REGION Network 15: EM - Abort Command
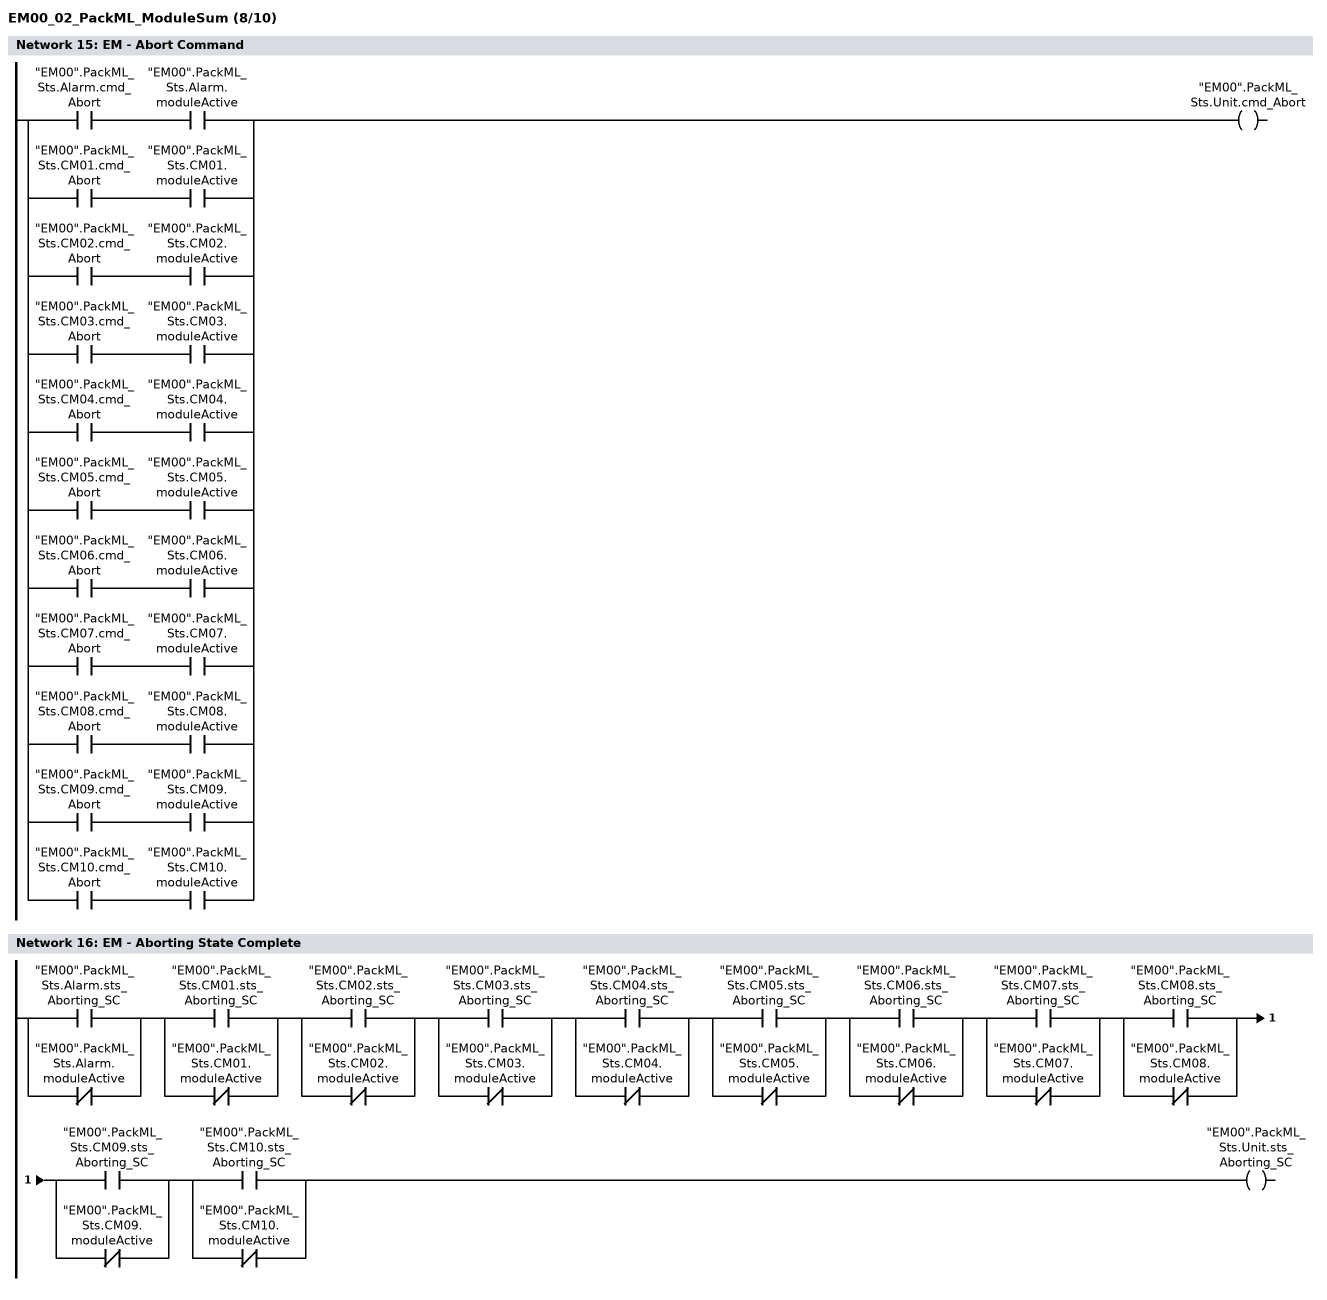
   RUNG wire#powerrail
      Contact( "EM00".PackML_Sts.Alarm.cmd_Abort )
      Contact( "EM00".PackML_Sts.Alarm.moduleActive )
      wire#w1
      Coil( "EM00".PackML_Sts.Unit.cmd_Abort )
   END_RUNG
   RUNG wire#powerrail
      Contact( "EM00".PackML_Sts.CM01.cmd_Abort )
      Contact( "EM00".PackML_Sts.CM01.moduleActive )
   END_RUNG wire#w1
   RUNG wire#powerrail
      Contact( "EM00".PackML_Sts.CM02.cmd_Abort )
      Contact( "EM00".PackML_Sts.CM02.moduleActive )
   END_RUNG wire#w1
   RUNG wire#powerrail
      Contact( "EM00".PackML_Sts.CM03.cmd_Abort )
      Contact( "EM00".PackML_Sts.CM03.moduleActive )
   END_RUNG wire#w1
   RUNG wire#powerrail
      Contact( "EM00".PackML_Sts.CM04.cmd_Abort )
      Contact( "EM00".PackML_Sts.CM04.moduleActive )
   END_RUNG wire#w1
   RUNG wire#powerrail
      Contact( "EM00".PackML_Sts.CM05.cmd_Abort )
      Contact( "EM00".PackML_Sts.CM05.moduleActive )
   END_RUNG wire#w1
   RUNG wire#powerrail
      Contact( "EM00".PackML_Sts.CM06.cmd_Abort )
      Contact( "EM00".PackML_Sts.CM06.moduleActive )
   END_RUNG wire#w1
   RUNG wire#powerrail
      Contact( "EM00".PackML_Sts.CM07.cmd_Abort )
      Contact( "EM00".PackML_Sts.CM07.moduleActive )
   END_RUNG wire#w1
   RUNG wire#powerrail
      Contact( "EM00".PackML_Sts.CM08.cmd_Abort )
      Contact( "EM00".PackML_Sts.CM08.moduleActive )
   END_RUNG wire#w1
   RUNG wire#powerrail
      Contact( "EM00".PackML_Sts.CM09.cmd_Abort )
      Contact( "EM00".PackML_Sts.CM09.moduleActive )
   END_RUNG wire#w1
   RUNG wire#powerrail
      Contact( "EM00".PackML_Sts.CM10.cmd_Abort )
      Contact( "EM00".PackML_Sts.CM10.moduleActive )
   END_RUNG wire#w1
   // the same network as SCL:
   "EM00".PackML_Sts.Unit.cmd_Abort := ("EM00".PackML_Sts.Alarm.cmd_Abort AND "EM00".PackML_Sts.Alarm.moduleActive) OR ("EM00".PackML_Sts.CM01.cmd_Abort AND "EM00".PackML_Sts.CM01.moduleActive) OR ("EM00".PackML_Sts.CM02.cmd_Abort AND "EM00".PackML_Sts.CM02.moduleActive) OR ("EM00".PackML_Sts.CM03.cmd_Abort AND "EM00".PackML_Sts.CM03.moduleActive) OR ("EM00".PackML_Sts.CM04.cmd_Abort AND "EM00".PackML_Sts.CM04.moduleActive) OR ("EM00".PackML_Sts.CM05.cmd_Abort AND "EM00".PackML_Sts.CM05.moduleActive) OR ("EM00".PackML_Sts.CM06.cmd_Abort AND "EM00".PackML_Sts.CM06.moduleActive) OR ("EM00".PackML_Sts.CM07.cmd_Abort AND "EM00".PackML_Sts.CM07.moduleActive) OR ("EM00".PackML_Sts.CM08.cmd_Abort AND "EM00".PackML_Sts.CM08.moduleActive) OR ("EM00".PackML_Sts.CM09.cmd_Abort AND "EM00".PackML_Sts.CM09.moduleActive) OR ("EM00".PackML_Sts.CM10.cmd_Abort AND "EM00".PackML_Sts.CM10.moduleActive);
END_REGION

REGION Network 16: EM - Aborting State Complete
   RUNG wire#powerrail
      Contact( "EM00".PackML_Sts.Alarm.sts_Aborting_SC )
      wire#w1
      Contact( "EM00".PackML_Sts.CM01.sts_Aborting_SC )
      wire#w2
      Contact( "EM00".PackML_Sts.CM02.sts_Aborting_SC )
      wire#w3
      Contact( "EM00".PackML_Sts.CM03.sts_Aborting_SC )
      wire#w4
      Contact( "EM00".PackML_Sts.CM04.sts_Aborting_SC )
      wire#w5
      Contact( "EM00".PackML_Sts.CM05.sts_Aborting_SC )
      wire#w6
      Contact( "EM00".PackML_Sts.CM06.sts_Aborting_SC )
      wire#w7
      Contact( "EM00".PackML_Sts.CM07.sts_Aborting_SC )
      wire#w8
      Contact( "EM00".PackML_Sts.CM08.sts_Aborting_SC )
      wire#w9
      Contact( "EM00".PackML_Sts.CM09.sts_Aborting_SC )
      wire#w10
      Contact( "EM00".PackML_Sts.CM10.sts_Aborting_SC )
      wire#w11
      Coil( "EM00".PackML_Sts.Unit.sts_Aborting_SC )
   END_RUNG
   RUNG wire#powerrail
      I_Contact( "EM00".PackML_Sts.Alarm.moduleActive )
   END_RUNG wire#w1
   RUNG wire#w1
      I_Contact( "EM00".PackML_Sts.CM01.moduleActive )
   END_RUNG wire#w2
   RUNG wire#w2
      I_Contact( "EM00".PackML_Sts.CM02.moduleActive )
   END_RUNG wire#w3
   RUNG wire#w3
      I_Contact( "EM00".PackML_Sts.CM03.moduleActive )
   END_RUNG wire#w4
   RUNG wire#w4
      I_Contact( "EM00".PackML_Sts.CM04.moduleActive )
   END_RUNG wire#w5
   RUNG wire#w5
      I_Contact( "EM00".PackML_Sts.CM05.moduleActive )
   END_RUNG wire#w6
   RUNG wire#w6
      I_Contact( "EM00".PackML_Sts.CM06.moduleActive )
   END_RUNG wire#w7
   RUNG wire#w7
      I_Contact( "EM00".PackML_Sts.CM07.moduleActive )
   END_RUNG wire#w8
   RUNG wire#w8
      I_Contact( "EM00".PackML_Sts.CM08.moduleActive )
   END_RUNG wire#w9
   RUNG wire#w9
      I_Contact( "EM00".PackML_Sts.CM09.moduleActive )
   END_RUNG wire#w10
   RUNG wire#w10
      I_Contact( "EM00".PackML_Sts.CM10.moduleActive )
   END_RUNG wire#w11
   // the same network as SCL:
   "EM00".PackML_Sts.Unit.sts_Aborting_SC := ("EM00".PackML_Sts.Alarm.sts_Aborting_SC OR NOT "EM00".PackML_Sts.Alarm.moduleActive) AND ("EM00".PackML_Sts.CM01.sts_Aborting_SC OR NOT "EM00".PackML_Sts.CM01.moduleActive) AND ("EM00".PackML_Sts.CM02.sts_Aborting_SC OR NOT "EM00".PackML_Sts.CM02.moduleActive) AND ("EM00".PackML_Sts.CM03.sts_Aborting_SC OR NOT "EM00".PackML_Sts.CM03.moduleActive) AND ("EM00".PackML_Sts.CM04.sts_Aborting_SC OR NOT "EM00".PackML_Sts.CM04.moduleActive) AND ("EM00".PackML_Sts.CM05.sts_Aborting_SC OR NOT "EM00".PackML_Sts.CM05.moduleActive) AND ("EM00".PackML_Sts.CM06.sts_Aborting_SC OR NOT "EM00".PackML_Sts.CM06.moduleActive) AND ("EM00".PackML_Sts.CM07.sts_Aborting_SC OR NOT "EM00".PackML_Sts.CM07.moduleActive) AND ("EM00".PackML_Sts.CM08.sts_Aborting_SC OR NOT "EM00".PackML_Sts.CM08.moduleActive) AND ("EM00".PackML_Sts.CM09.sts_Aborting_SC OR NOT "EM00".PackML_Sts.CM09.moduleActive) AND ("EM00".PackML_Sts.CM10.sts_Aborting_SC OR NOT "EM00".PackML_Sts.CM10.moduleActive);
END_REGION

REGION Network 17: EM - Clear Command
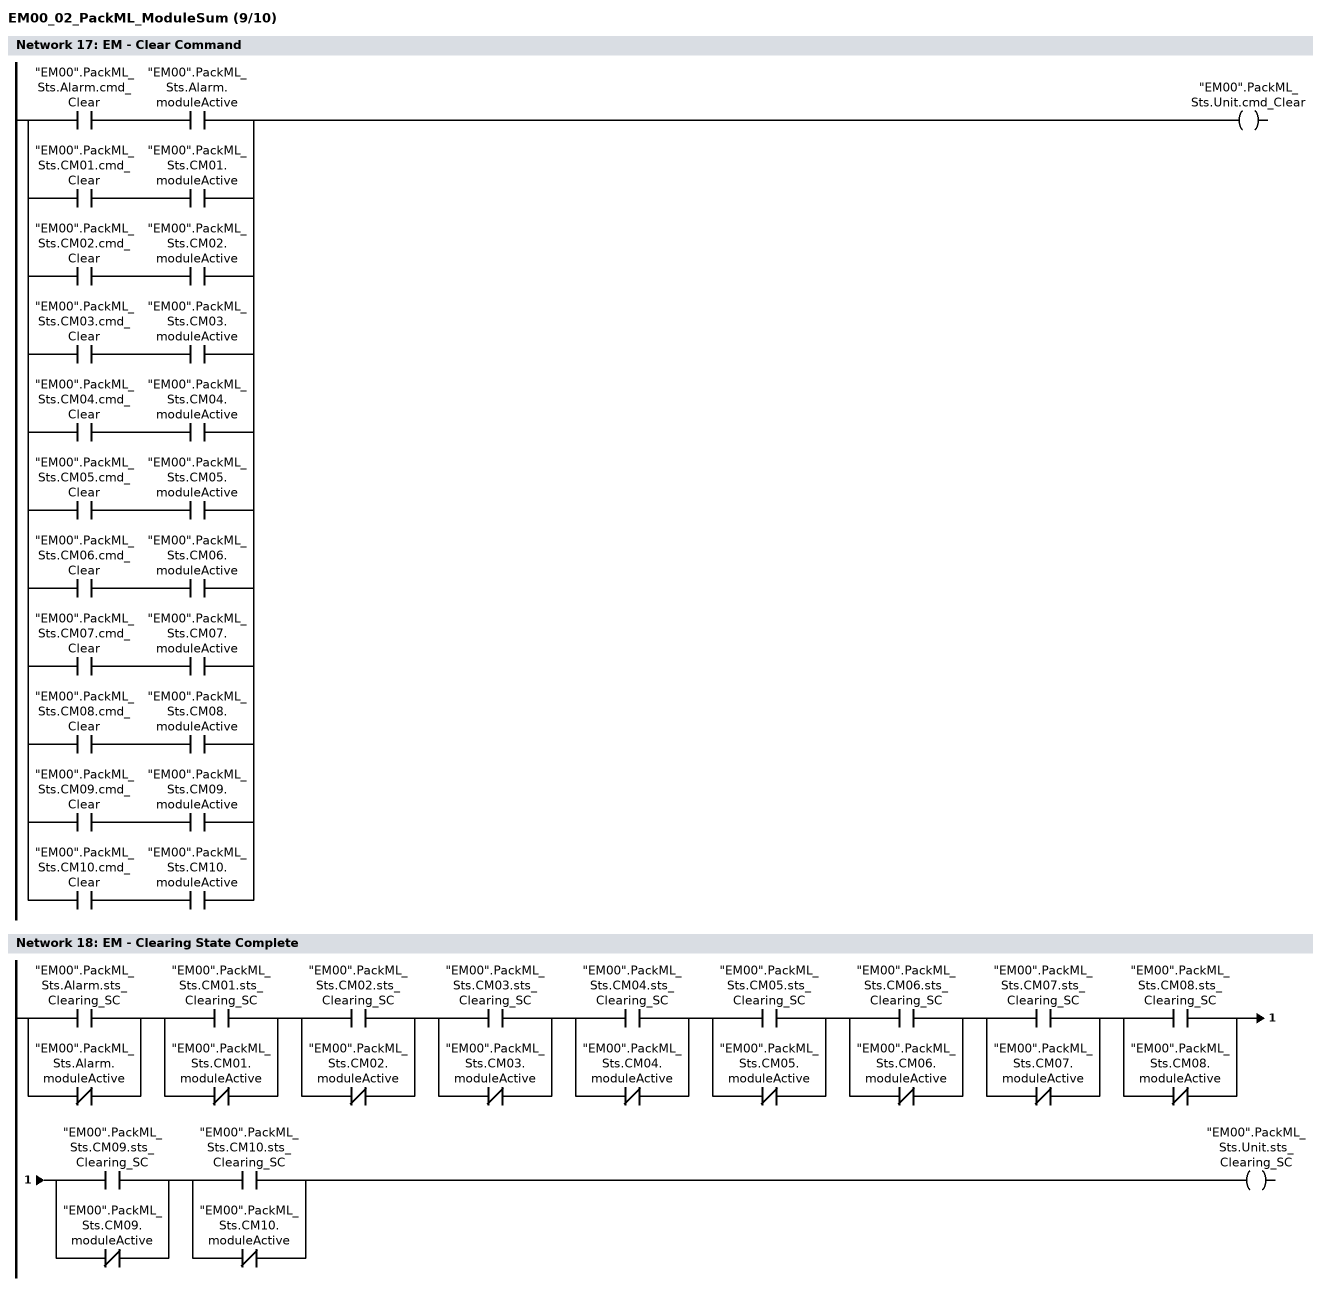
   RUNG wire#powerrail
      Contact( "EM00".PackML_Sts.Alarm.cmd_Clear )
      Contact( "EM00".PackML_Sts.Alarm.moduleActive )
      wire#w1
      Coil( "EM00".PackML_Sts.Unit.cmd_Clear )
   END_RUNG
   RUNG wire#powerrail
      Contact( "EM00".PackML_Sts.CM01.cmd_Clear )
      Contact( "EM00".PackML_Sts.CM01.moduleActive )
   END_RUNG wire#w1
   RUNG wire#powerrail
      Contact( "EM00".PackML_Sts.CM02.cmd_Clear )
      Contact( "EM00".PackML_Sts.CM02.moduleActive )
   END_RUNG wire#w1
   RUNG wire#powerrail
      Contact( "EM00".PackML_Sts.CM03.cmd_Clear )
      Contact( "EM00".PackML_Sts.CM03.moduleActive )
   END_RUNG wire#w1
   RUNG wire#powerrail
      Contact( "EM00".PackML_Sts.CM04.cmd_Clear )
      Contact( "EM00".PackML_Sts.CM04.moduleActive )
   END_RUNG wire#w1
   RUNG wire#powerrail
      Contact( "EM00".PackML_Sts.CM05.cmd_Clear )
      Contact( "EM00".PackML_Sts.CM05.moduleActive )
   END_RUNG wire#w1
   RUNG wire#powerrail
      Contact( "EM00".PackML_Sts.CM06.cmd_Clear )
      Contact( "EM00".PackML_Sts.CM06.moduleActive )
   END_RUNG wire#w1
   RUNG wire#powerrail
      Contact( "EM00".PackML_Sts.CM07.cmd_Clear )
      Contact( "EM00".PackML_Sts.CM07.moduleActive )
   END_RUNG wire#w1
   RUNG wire#powerrail
      Contact( "EM00".PackML_Sts.CM08.cmd_Clear )
      Contact( "EM00".PackML_Sts.CM08.moduleActive )
   END_RUNG wire#w1
   RUNG wire#powerrail
      Contact( "EM00".PackML_Sts.CM09.cmd_Clear )
      Contact( "EM00".PackML_Sts.CM09.moduleActive )
   END_RUNG wire#w1
   RUNG wire#powerrail
      Contact( "EM00".PackML_Sts.CM10.cmd_Clear )
      Contact( "EM00".PackML_Sts.CM10.moduleActive )
   END_RUNG wire#w1
   // the same network as SCL:
   "EM00".PackML_Sts.Unit.cmd_Clear := ("EM00".PackML_Sts.Alarm.cmd_Clear AND "EM00".PackML_Sts.Alarm.moduleActive) OR ("EM00".PackML_Sts.CM01.cmd_Clear AND "EM00".PackML_Sts.CM01.moduleActive) OR ("EM00".PackML_Sts.CM02.cmd_Clear AND "EM00".PackML_Sts.CM02.moduleActive) OR ("EM00".PackML_Sts.CM03.cmd_Clear AND "EM00".PackML_Sts.CM03.moduleActive) OR ("EM00".PackML_Sts.CM04.cmd_Clear AND "EM00".PackML_Sts.CM04.moduleActive) OR ("EM00".PackML_Sts.CM05.cmd_Clear AND "EM00".PackML_Sts.CM05.moduleActive) OR ("EM00".PackML_Sts.CM06.cmd_Clear AND "EM00".PackML_Sts.CM06.moduleActive) OR ("EM00".PackML_Sts.CM07.cmd_Clear AND "EM00".PackML_Sts.CM07.moduleActive) OR ("EM00".PackML_Sts.CM08.cmd_Clear AND "EM00".PackML_Sts.CM08.moduleActive) OR ("EM00".PackML_Sts.CM09.cmd_Clear AND "EM00".PackML_Sts.CM09.moduleActive) OR ("EM00".PackML_Sts.CM10.cmd_Clear AND "EM00".PackML_Sts.CM10.moduleActive);
END_REGION

REGION Network 18: EM - Clearing State Complete
   RUNG wire#powerrail
      Contact( "EM00".PackML_Sts.Alarm.sts_Clearing_SC )
      wire#w1
      Contact( "EM00".PackML_Sts.CM01.sts_Clearing_SC )
      wire#w2
      Contact( "EM00".PackML_Sts.CM02.sts_Clearing_SC )
      wire#w3
      Contact( "EM00".PackML_Sts.CM03.sts_Clearing_SC )
      wire#w4
      Contact( "EM00".PackML_Sts.CM04.sts_Clearing_SC )
      wire#w5
      Contact( "EM00".PackML_Sts.CM05.sts_Clearing_SC )
      wire#w6
      Contact( "EM00".PackML_Sts.CM06.sts_Clearing_SC )
      wire#w7
      Contact( "EM00".PackML_Sts.CM07.sts_Clearing_SC )
      wire#w8
      Contact( "EM00".PackML_Sts.CM08.sts_Clearing_SC )
      wire#w9
      Contact( "EM00".PackML_Sts.CM09.sts_Clearing_SC )
      wire#w10
      Contact( "EM00".PackML_Sts.CM10.sts_Clearing_SC )
      wire#w11
      Coil( "EM00".PackML_Sts.Unit.sts_Clearing_SC )
   END_RUNG
   RUNG wire#powerrail
      I_Contact( "EM00".PackML_Sts.Alarm.moduleActive )
   END_RUNG wire#w1
   RUNG wire#w1
      I_Contact( "EM00".PackML_Sts.CM01.moduleActive )
   END_RUNG wire#w2
   RUNG wire#w2
      I_Contact( "EM00".PackML_Sts.CM02.moduleActive )
   END_RUNG wire#w3
   RUNG wire#w3
      I_Contact( "EM00".PackML_Sts.CM03.moduleActive )
   END_RUNG wire#w4
   RUNG wire#w4
      I_Contact( "EM00".PackML_Sts.CM04.moduleActive )
   END_RUNG wire#w5
   RUNG wire#w5
      I_Contact( "EM00".PackML_Sts.CM05.moduleActive )
   END_RUNG wire#w6
   RUNG wire#w6
      I_Contact( "EM00".PackML_Sts.CM06.moduleActive )
   END_RUNG wire#w7
   RUNG wire#w7
      I_Contact( "EM00".PackML_Sts.CM07.moduleActive )
   END_RUNG wire#w8
   RUNG wire#w8
      I_Contact( "EM00".PackML_Sts.CM08.moduleActive )
   END_RUNG wire#w9
   RUNG wire#w9
      I_Contact( "EM00".PackML_Sts.CM09.moduleActive )
   END_RUNG wire#w10
   RUNG wire#w10
      I_Contact( "EM00".PackML_Sts.CM10.moduleActive )
   END_RUNG wire#w11
   // the same network as SCL:
   "EM00".PackML_Sts.Unit.sts_Clearing_SC := ("EM00".PackML_Sts.Alarm.sts_Clearing_SC OR NOT "EM00".PackML_Sts.Alarm.moduleActive) AND ("EM00".PackML_Sts.CM01.sts_Clearing_SC OR NOT "EM00".PackML_Sts.CM01.moduleActive) AND ("EM00".PackML_Sts.CM02.sts_Clearing_SC OR NOT "EM00".PackML_Sts.CM02.moduleActive) AND ("EM00".PackML_Sts.CM03.sts_Clearing_SC OR NOT "EM00".PackML_Sts.CM03.moduleActive) AND ("EM00".PackML_Sts.CM04.sts_Clearing_SC OR NOT "EM00".PackML_Sts.CM04.moduleActive) AND ("EM00".PackML_Sts.CM05.sts_Clearing_SC OR NOT "EM00".PackML_Sts.CM05.moduleActive) AND ("EM00".PackML_Sts.CM06.sts_Clearing_SC OR NOT "EM00".PackML_Sts.CM06.moduleActive) AND ("EM00".PackML_Sts.CM07.sts_Clearing_SC OR NOT "EM00".PackML_Sts.CM07.moduleActive) AND ("EM00".PackML_Sts.CM08.sts_Clearing_SC OR NOT "EM00".PackML_Sts.CM08.moduleActive) AND ("EM00".PackML_Sts.CM09.sts_Clearing_SC OR NOT "EM00".PackML_Sts.CM09.moduleActive) AND ("EM00".PackML_Sts.CM10.sts_Clearing_SC OR NOT "EM00".PackML_Sts.CM10.moduleActive);
END_REGION

REGION Network 19: EM - Execute State Complete
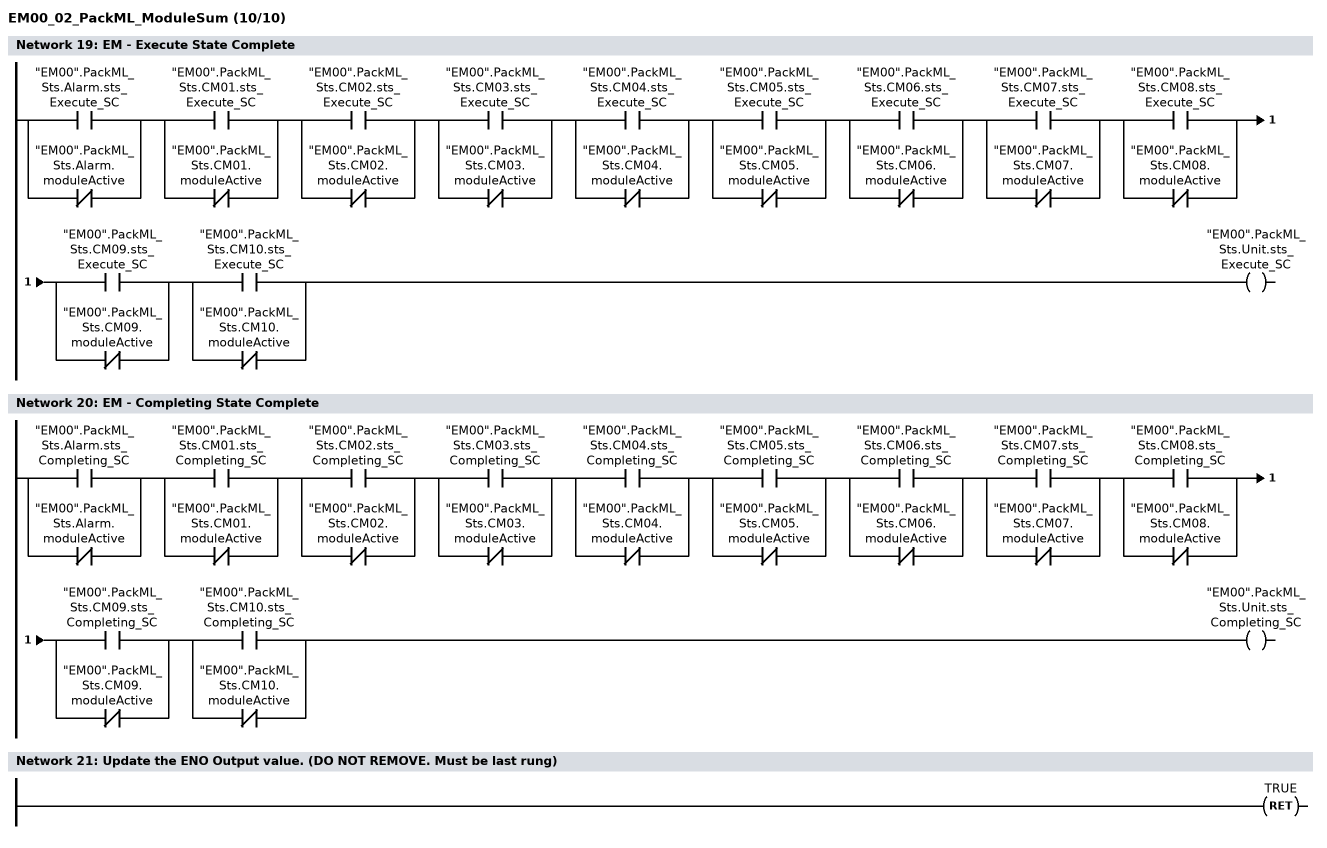
   RUNG wire#powerrail
      Contact( "EM00".PackML_Sts.Alarm.sts_Execute_SC )
      wire#w1
      Contact( "EM00".PackML_Sts.CM01.sts_Execute_SC )
      wire#w2
      Contact( "EM00".PackML_Sts.CM02.sts_Execute_SC )
      wire#w3
      Contact( "EM00".PackML_Sts.CM03.sts_Execute_SC )
      wire#w4
      Contact( "EM00".PackML_Sts.CM04.sts_Execute_SC )
      wire#w5
      Contact( "EM00".PackML_Sts.CM05.sts_Execute_SC )
      wire#w6
      Contact( "EM00".PackML_Sts.CM06.sts_Execute_SC )
      wire#w7
      Contact( "EM00".PackML_Sts.CM07.sts_Execute_SC )
      wire#w8
      Contact( "EM00".PackML_Sts.CM08.sts_Execute_SC )
      wire#w9
      Contact( "EM00".PackML_Sts.CM09.sts_Execute_SC )
      wire#w10
      Contact( "EM00".PackML_Sts.CM10.sts_Execute_SC )
      wire#w11
      Coil( "EM00".PackML_Sts.Unit.sts_Execute_SC )
   END_RUNG
   RUNG wire#powerrail
      I_Contact( "EM00".PackML_Sts.Alarm.moduleActive )
   END_RUNG wire#w1
   RUNG wire#w1
      I_Contact( "EM00".PackML_Sts.CM01.moduleActive )
   END_RUNG wire#w2
   RUNG wire#w2
      I_Contact( "EM00".PackML_Sts.CM02.moduleActive )
   END_RUNG wire#w3
   RUNG wire#w3
      I_Contact( "EM00".PackML_Sts.CM03.moduleActive )
   END_RUNG wire#w4
   RUNG wire#w4
      I_Contact( "EM00".PackML_Sts.CM04.moduleActive )
   END_RUNG wire#w5
   RUNG wire#w5
      I_Contact( "EM00".PackML_Sts.CM05.moduleActive )
   END_RUNG wire#w6
   RUNG wire#w6
      I_Contact( "EM00".PackML_Sts.CM06.moduleActive )
   END_RUNG wire#w7
   RUNG wire#w7
      I_Contact( "EM00".PackML_Sts.CM07.moduleActive )
   END_RUNG wire#w8
   RUNG wire#w8
      I_Contact( "EM00".PackML_Sts.CM08.moduleActive )
   END_RUNG wire#w9
   RUNG wire#w9
      I_Contact( "EM00".PackML_Sts.CM09.moduleActive )
   END_RUNG wire#w10
   RUNG wire#w10
      I_Contact( "EM00".PackML_Sts.CM10.moduleActive )
   END_RUNG wire#w11
   // the same network as SCL:
   "EM00".PackML_Sts.Unit.sts_Execute_SC := ("EM00".PackML_Sts.Alarm.sts_Execute_SC OR NOT "EM00".PackML_Sts.Alarm.moduleActive) AND ("EM00".PackML_Sts.CM01.sts_Execute_SC OR NOT "EM00".PackML_Sts.CM01.moduleActive) AND ("EM00".PackML_Sts.CM02.sts_Execute_SC OR NOT "EM00".PackML_Sts.CM02.moduleActive) AND ("EM00".PackML_Sts.CM03.sts_Execute_SC OR NOT "EM00".PackML_Sts.CM03.moduleActive) AND ("EM00".PackML_Sts.CM04.sts_Execute_SC OR NOT "EM00".PackML_Sts.CM04.moduleActive) AND ("EM00".PackML_Sts.CM05.sts_Execute_SC OR NOT "EM00".PackML_Sts.CM05.moduleActive) AND ("EM00".PackML_Sts.CM06.sts_Execute_SC OR NOT "EM00".PackML_Sts.CM06.moduleActive) AND ("EM00".PackML_Sts.CM07.sts_Execute_SC OR NOT "EM00".PackML_Sts.CM07.moduleActive) AND ("EM00".PackML_Sts.CM08.sts_Execute_SC OR NOT "EM00".PackML_Sts.CM08.moduleActive) AND ("EM00".PackML_Sts.CM09.sts_Execute_SC OR NOT "EM00".PackML_Sts.CM09.moduleActive) AND ("EM00".PackML_Sts.CM10.sts_Execute_SC OR NOT "EM00".PackML_Sts.CM10.moduleActive);
END_REGION

REGION Network 20: EM - Completing State Complete
   RUNG wire#powerrail
      Contact( "EM00".PackML_Sts.Alarm.sts_Completing_SC )
      wire#w1
      Contact( "EM00".PackML_Sts.CM01.sts_Completing_SC )
      wire#w2
      Contact( "EM00".PackML_Sts.CM02.sts_Completing_SC )
      wire#w3
      Contact( "EM00".PackML_Sts.CM03.sts_Completing_SC )
      wire#w4
      Contact( "EM00".PackML_Sts.CM04.sts_Completing_SC )
      wire#w5
      Contact( "EM00".PackML_Sts.CM05.sts_Completing_SC )
      wire#w6
      Contact( "EM00".PackML_Sts.CM06.sts_Completing_SC )
      wire#w7
      Contact( "EM00".PackML_Sts.CM07.sts_Completing_SC )
      wire#w8
      Contact( "EM00".PackML_Sts.CM08.sts_Completing_SC )
      wire#w9
      Contact( "EM00".PackML_Sts.CM09.sts_Completing_SC )
      wire#w10
      Contact( "EM00".PackML_Sts.CM10.sts_Completing_SC )
      wire#w11
      Coil( "EM00".PackML_Sts.Unit.sts_Completing_SC )
   END_RUNG
   RUNG wire#powerrail
      I_Contact( "EM00".PackML_Sts.Alarm.moduleActive )
   END_RUNG wire#w1
   RUNG wire#w1
      I_Contact( "EM00".PackML_Sts.CM01.moduleActive )
   END_RUNG wire#w2
   RUNG wire#w2
      I_Contact( "EM00".PackML_Sts.CM02.moduleActive )
   END_RUNG wire#w3
   RUNG wire#w3
      I_Contact( "EM00".PackML_Sts.CM03.moduleActive )
   END_RUNG wire#w4
   RUNG wire#w4
      I_Contact( "EM00".PackML_Sts.CM04.moduleActive )
   END_RUNG wire#w5
   RUNG wire#w5
      I_Contact( "EM00".PackML_Sts.CM05.moduleActive )
   END_RUNG wire#w6
   RUNG wire#w6
      I_Contact( "EM00".PackML_Sts.CM06.moduleActive )
   END_RUNG wire#w7
   RUNG wire#w7
      I_Contact( "EM00".PackML_Sts.CM07.moduleActive )
   END_RUNG wire#w8
   RUNG wire#w8
      I_Contact( "EM00".PackML_Sts.CM08.moduleActive )
   END_RUNG wire#w9
   RUNG wire#w9
      I_Contact( "EM00".PackML_Sts.CM09.moduleActive )
   END_RUNG wire#w10
   RUNG wire#w10
      I_Contact( "EM00".PackML_Sts.CM10.moduleActive )
   END_RUNG wire#w11
   // the same network as SCL:
   "EM00".PackML_Sts.Unit.sts_Completing_SC := ("EM00".PackML_Sts.Alarm.sts_Completing_SC OR NOT "EM00".PackML_Sts.Alarm.moduleActive) AND ("EM00".PackML_Sts.CM01.sts_Completing_SC OR NOT "EM00".PackML_Sts.CM01.moduleActive) AND ("EM00".PackML_Sts.CM02.sts_Completing_SC OR NOT "EM00".PackML_Sts.CM02.moduleActive) AND ("EM00".PackML_Sts.CM03.sts_Completing_SC OR NOT "EM00".PackML_Sts.CM03.moduleActive) AND ("EM00".PackML_Sts.CM04.sts_Completing_SC OR NOT "EM00".PackML_Sts.CM04.moduleActive) AND ("EM00".PackML_Sts.CM05.sts_Completing_SC OR NOT "EM00".PackML_Sts.CM05.moduleActive) AND ("EM00".PackML_Sts.CM06.sts_Completing_SC OR NOT "EM00".PackML_Sts.CM06.moduleActive) AND ("EM00".PackML_Sts.CM07.sts_Completing_SC OR NOT "EM00".PackML_Sts.CM07.moduleActive) AND ("EM00".PackML_Sts.CM08.sts_Completing_SC OR NOT "EM00".PackML_Sts.CM08.moduleActive) AND ("EM00".PackML_Sts.CM09.sts_Completing_SC OR NOT "EM00".PackML_Sts.CM09.moduleActive) AND ("EM00".PackML_Sts.CM10.sts_Completing_SC OR NOT "EM00".PackML_Sts.CM10.moduleActive);
END_REGION

REGION Network 21: Update the ENO Output value. (DO NOT REMOVE. Must be last rung)
   RUNG wire#powerrail
      ReturnCoil( TRUE )
   END_RUNG
   // the same network as SCL:
   ENO := TRUE;
   RETURN;
END_REGION
END_FUNCTION_BLOCK

FUNCTION_BLOCK "EM00_CM01_MainOpStation"   // FB31651, LAD
TITLE = EM00_CM01_MainOpStation
{ S7_Optimized_Access := 'TRUE' }
AUTHOR : tech.team.motioncontrol@siemens.com
FAMILY : CPG
VERSION : 1.1
// Support: tech.team.motioncontrol@siemens.com
   VAR
      instAlarm_EStop : "CPG_Event";   // Alarm Event - EStop pressed (Event instance)
      instAlarm_HMI_StopPB : "CPG_Event";   // Alarm Event - HMI Stop PB pressed (Event instance)
      instStatus_WaitingForStartCmd : "CPG_Event";   // Status Event - waiting for start command (Event instance)
      instStatus_WaitingForResetCmd : "CPG_Event";   // Status Event - waiting for reset command (Event instance)
      instAlarm_Hold_PB : "CPG_Event";   // Alarm Event - HMI Held PB pressed (Event instance)
      instStatus_WaitingForUnHoldCmd : "CPG_Event";   // Status Event - waiting for unhold command (Event instance)
      instTimer_StartingDelay_SC : IEC_TIMER;   // IEC Timer - starting delay (demo only - used to slow state model transition)
      instTimer_CompletingDelay_SC : IEC_TIMER;   // IEC Timer - completing delay (demo only - used to slow state model transition)
      instTimer_AbortingDelay_SC : IEC_TIMER;   // IEC Timer - aborting delay (demo only - used to slow state model transition)
      instTimer_StoppingDelay_SC : IEC_TIMER;   // IEC Timer - stopping delay (demo only - used to slow state model transition)
      instTimer_ResettingDelay_SC : IEC_TIMER;   // IEC Timer - resetting delay (demo only - used to slow state model transition)
      instTimer_HoldingDelay_SC : IEC_TIMER;   // IEC Timer - holding delay (demo only - used to slow state model transition)
      instTimer_UnHoldingDelay_SC : IEC_TIMER;   // IEC Timer - un-holding delay (demo only - used to slow state model transition)
      instTimer_SuspendingDelay_SC : IEC_TIMER;   // IEC Timer - suspending delay (demo only - used to slow state model transition)
      instTimer_UnSuspendingDelay_SC : IEC_TIMER;   // IEC Timer - un-suspending delay (demo only - used to slow state model transition)
      instTimer_ClearingDelay_SC : IEC_TIMER;   // IEC Timer - clearing delay (demo only - used to slow state model transition)
      FTriggerTest_Instance : "FTriggerTest";
   END_VAR
BEGIN

REGION Network 1: *** Begin the Setpoint Management Information Section ***
END_REGION

REGION Network 2: *** Begin the Logic Section ***
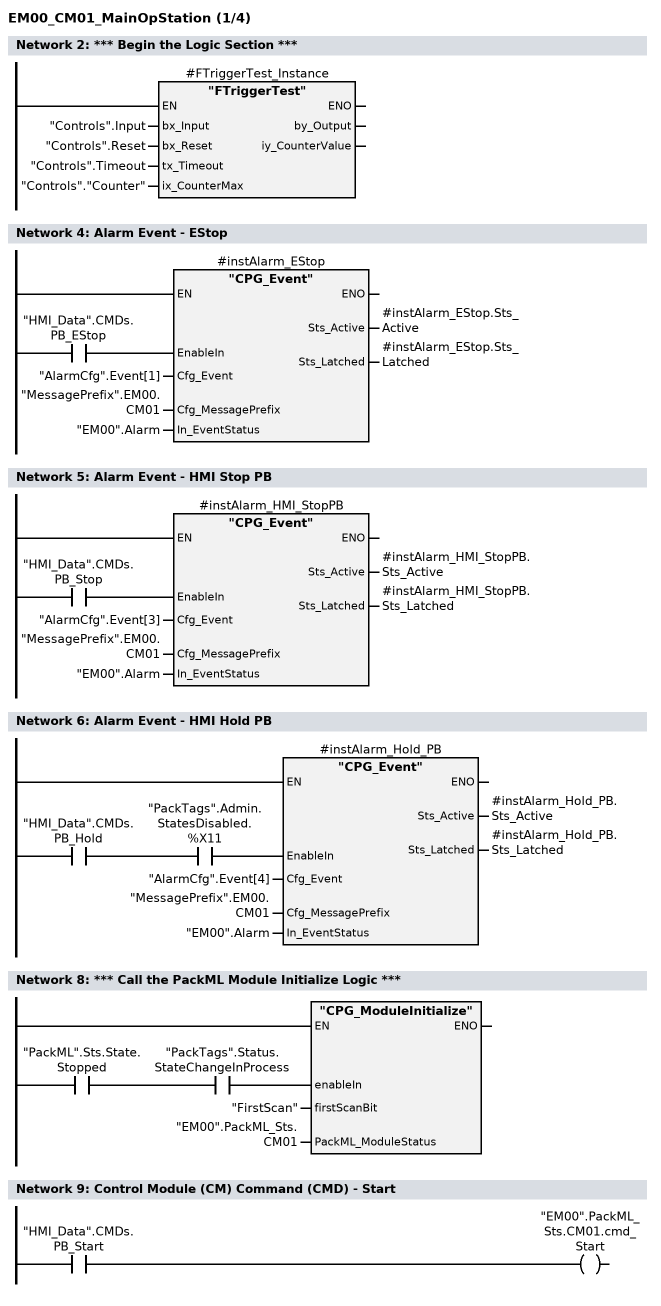
   RUNG wire#powerrail
      #FTriggerTest_Instance(bx_Input := "Controls".Input, bx_Reset := "Controls".Reset, tx_Timeout := "Controls".Timeout, ix_CounterMax := "Controls"."Counter", by_Output =>, iy_CounterValue =>)
   END_RUNG
   // the same network as SCL:
   #FTriggerTest_Instance(bx_Input := "Controls".Input,   // "FTriggerTest"
                          bx_Reset := "Controls".Reset,
                          tx_Timeout := "Controls".Timeout,
                          ix_CounterMax := "Controls"."Counter");
END_REGION

REGION Network 3: *** Begin the Event Information Section ***
END_REGION

REGION Network 4: Alarm Event - EStop
   RUNG wire#powerrail
      #instAlarm_EStop(EnableIn := wire#w1, Cfg_Event := "AlarmCfg".Event[1], Cfg_MessagePrefix := "MessagePrefix".EM00.CM01, In_EventStatus := "EM00".Alarm, Sts_Active => #instAlarm_EStop.Sts_Active, Sts_Latched => #instAlarm_EStop.Sts_Latched)
   END_RUNG
   RUNG wire#powerrail
      Contact( "HMI_Data".CMDs.PB_EStop )
   END_RUNG wire#w1
   // the same network as SCL:
   #instAlarm_EStop(EnableIn := "HMI_Data".CMDs.PB_EStop,   // "CPG_Event"
                    Cfg_Event := "AlarmCfg".Event[1],
                    Cfg_MessagePrefix := "MessagePrefix".EM00.CM01,
                    In_EventStatus := "EM00".Alarm,
                    Sts_Active => #instAlarm_EStop.Sts_Active,
                    Sts_Latched => #instAlarm_EStop.Sts_Latched);
END_REGION

REGION Network 5: Alarm Event - HMI Stop PB
   RUNG wire#powerrail
      #instAlarm_HMI_StopPB(EnableIn := wire#w1, Cfg_Event := "AlarmCfg".Event[3], Cfg_MessagePrefix := "MessagePrefix".EM00.CM01, In_EventStatus := "EM00".Alarm, Sts_Active => #instAlarm_HMI_StopPB.Sts_Active, Sts_Latched => #instAlarm_HMI_StopPB.Sts_Latched)
   END_RUNG
   RUNG wire#powerrail
      Contact( "HMI_Data".CMDs.PB_Stop )
   END_RUNG wire#w1
   // the same network as SCL:
   #instAlarm_HMI_StopPB(EnableIn := "HMI_Data".CMDs.PB_Stop,   // "CPG_Event"
                         Cfg_Event := "AlarmCfg".Event[3],
                         Cfg_MessagePrefix := "MessagePrefix".EM00.CM01,
                         In_EventStatus := "EM00".Alarm,
                         Sts_Active => #instAlarm_HMI_StopPB.Sts_Active,
                         Sts_Latched => #instAlarm_HMI_StopPB.Sts_Latched);
END_REGION

REGION Network 6: Alarm Event - HMI Hold PB
   RUNG wire#powerrail
      #instAlarm_Hold_PB(EnableIn := wire#w1, Cfg_Event := "AlarmCfg".Event[4], Cfg_MessagePrefix := "MessagePrefix".EM00.CM01, In_EventStatus := "EM00".Alarm, Sts_Active => #instAlarm_Hold_PB.Sts_Active, Sts_Latched => #instAlarm_Hold_PB.Sts_Latched)
   END_RUNG
   RUNG wire#powerrail
      Contact( "HMI_Data".CMDs.PB_Hold )
      Contact( "PackTags".Admin.StatesDisabled.%X11 )
   END_RUNG wire#w1
   // the same network as SCL:
   #instAlarm_Hold_PB(EnableIn := "HMI_Data".CMDs.PB_Hold AND "PackTags".Admin.StatesDisabled.%X11,   // "CPG_Event"
                      Cfg_Event := "AlarmCfg".Event[4],
                      Cfg_MessagePrefix := "MessagePrefix".EM00.CM01,
                      In_EventStatus := "EM00".Alarm,
                      Sts_Active => #instAlarm_Hold_PB.Sts_Active,
                      Sts_Latched => #instAlarm_Hold_PB.Sts_Latched);
END_REGION

REGION Network 7: *** Begin the State Model Status Feedback Section ***
END_REGION

REGION Network 8: *** Call the PackML Module Initialize Logic ***
   RUNG wire#powerrail
      "CPG_ModuleInitialize"(enableIn := wire#w1, firstScanBit := "FirstScan", PackML_ModuleStatus := "EM00".PackML_Sts.CM01)
   END_RUNG
   RUNG wire#powerrail
      Contact( "PackML".Sts.State.Stopped )
      Contact( "PackTags".Status.StateChangeInProcess )
   END_RUNG wire#w1
   // the same network as SCL:
   "CPG_ModuleInitialize"(enableIn := "PackML".Sts.State.Stopped AND "PackTags".Status.StateChangeInProcess,
                          firstScanBit := "FirstScan",
                          PackML_ModuleStatus := "EM00".PackML_Sts.CM01);
END_REGION

REGION Network 9: Control Module (CM) Command (CMD) - Start
   RUNG wire#powerrail
      Contact( "HMI_Data".CMDs.PB_Start )
      Coil( "EM00".PackML_Sts.CM01.cmd_Start )
   END_RUNG
   // the same network as SCL:
   "EM00".PackML_Sts.CM01.cmd_Start := "HMI_Data".CMDs.PB_Start;
END_REGION

REGION Network 10: Status Event message for HMI - Waiting for Start PB